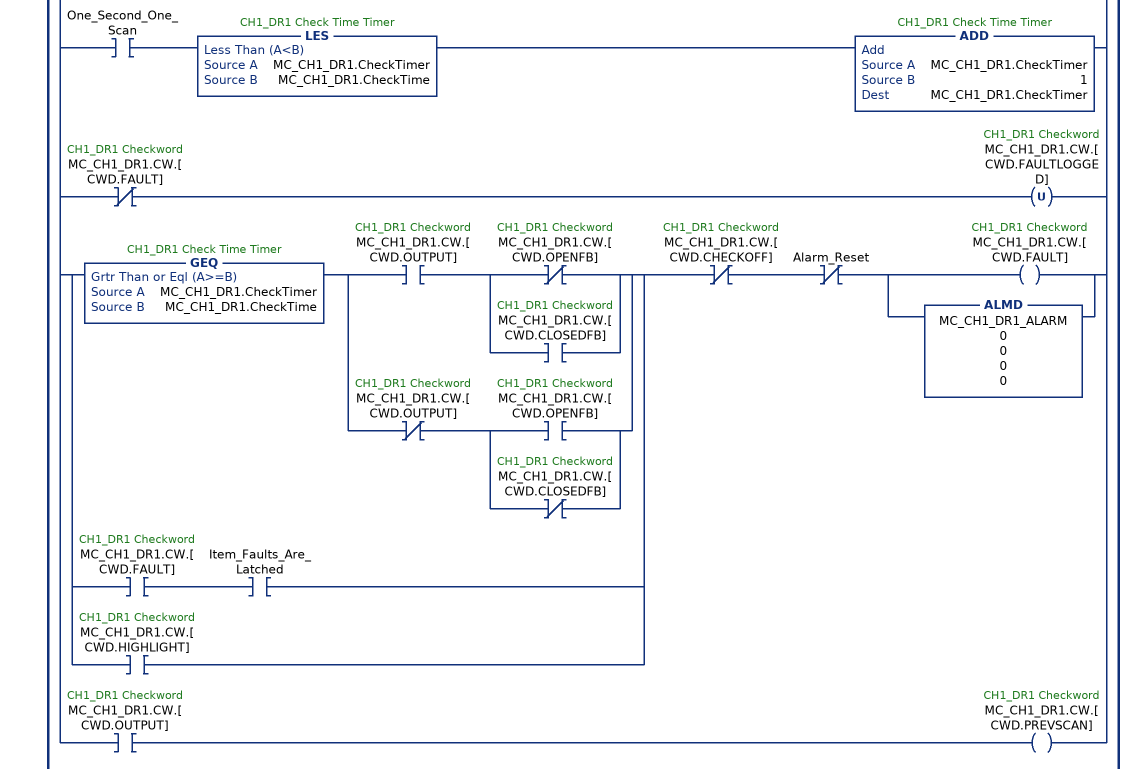
   14: [NEQ(MC_CH1_DR1.DriveBits,0) OTE(MC_CH1_DR1.CW.[CWD.AUTODRV]) ,[XIC(MC_CH1_DR1.CW.[CWD.AUTODRV]) XIO(MC_CH1_DR1.CW.[CWD.MANUAL]) ,XIC(MC_CH1_DR1.CW.[CWD.MANDRV]) XIC(MC_CH1_DR1.CW.[CWD.MANUAL]) ] OTE(MC_CH1_DR1.CW.[CWD.OUTPUT]) ,XIC(MC_CH1_DR1.CW.[CWD.OUTPUT]) OTE(MC_CH1_DR1_DR) ,XIC(S:FS) [OTU(MC_CH1_DR1.CW.[CWD.MANUAL]) ,LEQ(MC_CH1_DR1.CheckTime,0) MOV(Default_Check_Time,MC_CH1_DR1.CheckTime) ] ,[[XIC(MC_CH1_DR1_O) XIO(Item_Simulation_Flag) ,XIC(Item_Simulation_Flag) XIC(MC_CH1_DR1.CW.[CWD.OUTPUT]) XIO(MC_CH1_DR1.CW.[CWD.SIMFAIL]) ] OTE(MC_CH1_DR1.CW.[CWD.OPENFB]) ,[XIC(MC_CH1_DR1_C) XIO(Item_Simulation_Flag) ,XIC(Item_Simulation_Flag) XIO(MC_CH1_DR1.CW.[CWD.OUTPUT]) XIO(MC_CH1_DR1.CW.[CWD.SIMFAIL]) ] OTE(MC_CH1_DR1.CW.[CWD.CLOSEDFB]) ] ,[XIC(MC_CH1_DR1.CW.[CWD.OUTPUT]) XIO(MC_CH1_DR1.CW.[CWD.PREVSCAN]) ,XIO(MC_CH1_DR1.CW.[CWD.OUTPUT]) XIC(MC_CH1_DR1.CW.[CWD.PREVSCAN]) ] CLR(MC_CH1_DR1.CheckTimer) ,XIC(One_Second_One_Scan) LES(MC_CH1_DR1.CheckTimer,MC_CH1_DR1.CheckTime) ADD(MC_CH1_DR1.CheckTimer,1,MC_CH1_DR1.CheckTimer) ,XIO(MC_CH1_DR1.CW.[CWD.FAULT]) OTU(MC_CH1_DR1.CW.[CWD.FAULTLOGGED]) ,[GEQ(MC_CH1_DR1.CheckTimer,MC_CH1_DR1.CheckTime) [XIC(MC_CH1_DR1.CW.[CWD.OUTPUT]) [XIO(MC_CH1_DR1.CW.[CWD.OPENFB]) ,XIC(MC_CH1_DR1.CW.[CWD.CLOSEDFB]) ] ,XIO(MC_CH1_DR1.CW.[CWD.OUTPUT]) [XIC(MC_CH1_DR1.CW.[CWD.OPENFB]) ,XIO(MC_CH1_DR1.CW.[CWD.CLOSEDFB]) ] ] ,XIC(MC_CH1_DR1.CW.[CWD.FAULT]) XIC(Item_Faults_Are_Latched) ,XIC(MC_CH1_DR1.CW.[CWD.HIGHLIGHT]) ] XIO(MC_CH1_DR1.CW.[CWD.CHECKOFF]) XIO(Alarm_Reset) [OTE(MC_CH1_DR1.CW.[CWD.FAULT]) ,ALMD(MC_CH1_DR1_ALARM,0,0,0,0) ] ,XIC(MC_CH1_DR1.CW.[CWD.OUTPUT]) OTE(MC_CH1_DR1.CW.[CWD.PREVSCAN]) ];
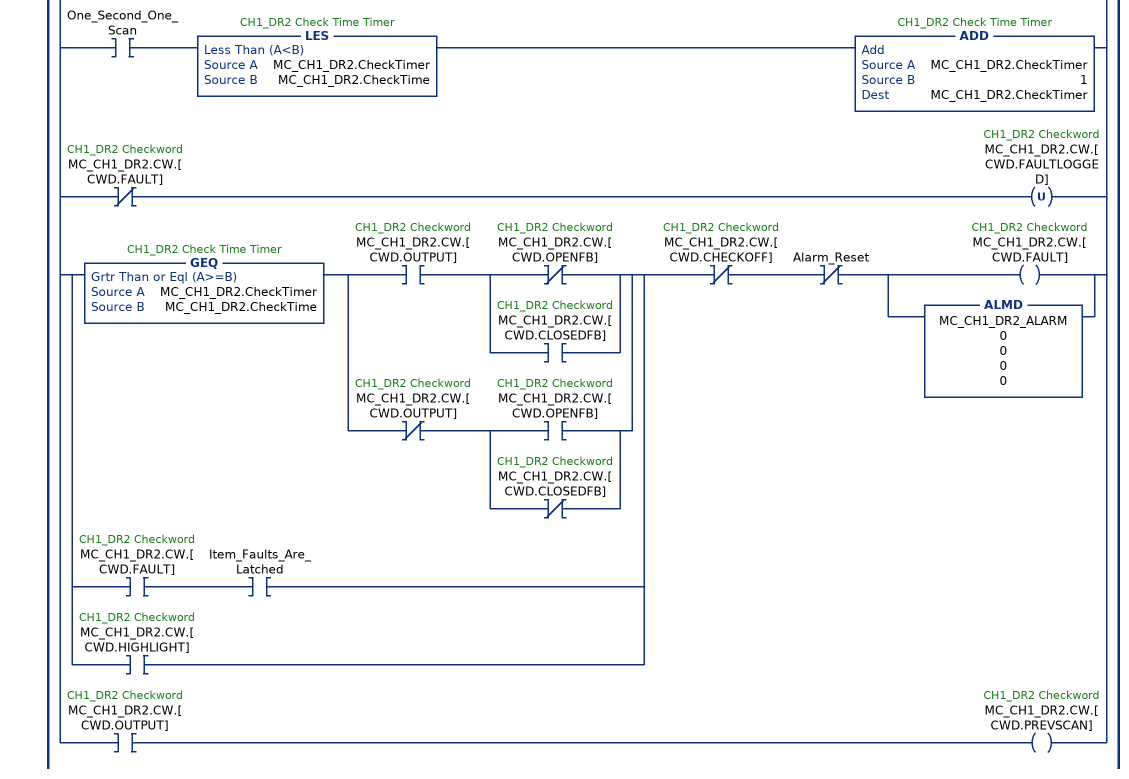
   15: [NEQ(MC_CH1_DR2.DriveBits,0) OTE(MC_CH1_DR2.CW.[CWD.AUTODRV]) ,[XIC(MC_CH1_DR2.CW.[CWD.AUTODRV]) XIO(MC_CH1_DR2.CW.[CWD.MANUAL]) ,XIC(MC_CH1_DR2.CW.[CWD.MANDRV]) XIC(MC_CH1_DR2.CW.[CWD.MANUAL]) ] OTE(MC_CH1_DR2.CW.[CWD.OUTPUT]) ,XIC(MC_CH1_DR2.CW.[CWD.OUTPUT]) OTE(MC_CH1_DR2_DR) ,XIC(S:FS) [OTU(MC_CH1_DR2.CW.[CWD.MANUAL]) ,LEQ(MC_CH1_DR2.CheckTime,0) MOV(Default_Check_Time,MC_CH1_DR2.CheckTime) ] ,[[XIC(MC_CH1_DR2_O) XIO(Item_Simulation_Flag) ,XIC(Item_Simulation_Flag) XIC(MC_CH1_DR2.CW.[CWD.OUTPUT]) XIO(MC_CH1_DR2.CW.[CWD.SIMFAIL]) ] OTE(MC_CH1_DR2.CW.[CWD.OPENFB]) ,[XIC(MC_CH1_DR2_C) XIO(Item_Simulation_Flag) ,XIC(Item_Simulation_Flag) XIO(MC_CH1_DR2.CW.[CWD.OUTPUT]) XIO(MC_CH1_DR2.CW.[CWD.SIMFAIL]) ] OTE(MC_CH1_DR2.CW.[CWD.CLOSEDFB]) ] ,[XIC(MC_CH1_DR2.CW.[CWD.OUTPUT]) XIO(MC_CH1_DR2.CW.[CWD.PREVSCAN]) ,XIO(MC_CH1_DR2.CW.[CWD.OUTPUT]) XIC(MC_CH1_DR2.CW.[CWD.PREVSCAN]) ] CLR(MC_CH1_DR2.CheckTimer) ,XIC(One_Second_One_Scan) LES(MC_CH1_DR2.CheckTimer,MC_CH1_DR2.CheckTime) ADD(MC_CH1_DR2.CheckTimer,1,MC_CH1_DR2.CheckTimer) ,XIO(MC_CH1_DR2.CW.[CWD.FAULT]) OTU(MC_CH1_DR2.CW.[CWD.FAULTLOGGED]) ,[GEQ(MC_CH1_DR2.CheckTimer,MC_CH1_DR2.CheckTime) [XIC(MC_CH1_DR2.CW.[CWD.OUTPUT]) [XIO(MC_CH1_DR2.CW.[CWD.OPENFB]) ,XIC(MC_CH1_DR2.CW.[CWD.CLOSEDFB]) ] ,XIO(MC_CH1_DR2.CW.[CWD.OUTPUT]) [XIC(MC_CH1_DR2.CW.[CWD.OPENFB]) ,XIO(MC_CH1_DR2.CW.[CWD.CLOSEDFB]) ] ] ,XIC(MC_CH1_DR2.CW.[CWD.FAULT]) XIC(Item_Faults_Are_Latched) ,XIC(MC_CH1_DR2.CW.[CWD.HIGHLIGHT]) ] XIO(MC_CH1_DR2.CW.[CWD.CHECKOFF]) XIO(Alarm_Reset) [OTE(MC_CH1_DR2.CW.[CWD.FAULT]) ,ALMD(MC_CH1_DR2_ALARM,0,0,0,0) ] ,XIC(MC_CH1_DR2.CW.[CWD.OUTPUT]) OTE(MC_CH1_DR2.CW.[CWD.PREVSCAN]) ];
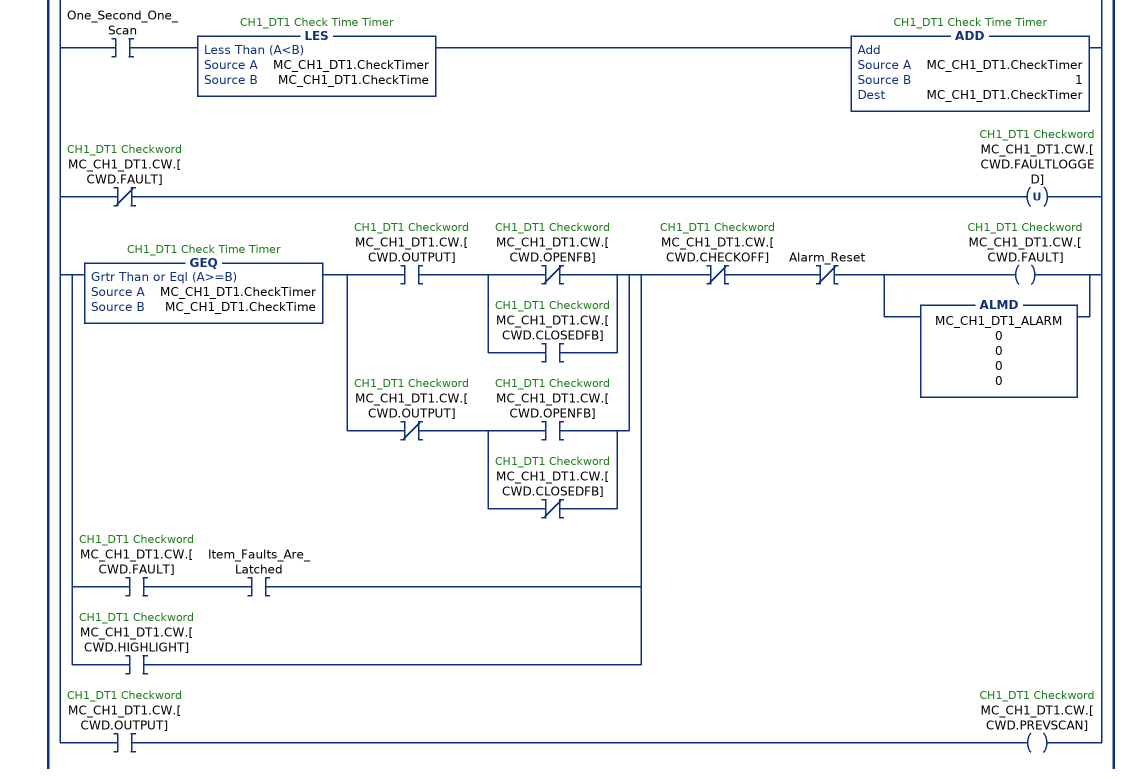
   16: [NEQ(MC_CH1_DT1.DriveBits,0) OTE(MC_CH1_DT1.CW.[CWD.AUTODRV]) ,[XIC(MC_CH1_DT1.CW.[CWD.AUTODRV]) XIO(MC_CH1_DT1.CW.[CWD.MANUAL]) ,XIC(MC_CH1_DT1.CW.[CWD.MANDRV]) XIC(MC_CH1_DT1.CW.[CWD.MANUAL]) ] OTE(MC_CH1_DT1.CW.[CWD.OUTPUT]) ,XIC(MC_CH1_DT1.CW.[CWD.OUTPUT]) OTE(MC_CH1_DT1_DR) ,XIC(S:FS) [OTU(MC_CH1_DT1.CW.[CWD.MANUAL]) ,LEQ(MC_CH1_DT1.CheckTime,0) MOV(Default_Check_Time,MC_CH1_DT1.CheckTime) ] ,[[XIC(MC_CH1_DT1_O) XIO(Item_Simulation_Flag) ,XIC(Item_Simulation_Flag) XIC(MC_CH1_DT1.CW.[CWD.OUTPUT]) XIO(MC_CH1_DT1.CW.[CWD.SIMFAIL]) ] OTE(MC_CH1_DT1.CW.[CWD.OPENFB]) ,[XIC(MC_CH1_DT1_C) XIO(Item_Simulation_Flag) ,XIC(Item_Simulation_Flag) XIO(MC_CH1_DT1.CW.[CWD.OUTPUT]) XIO(MC_CH1_DT1.CW.[CWD.SIMFAIL]) ] OTE(MC_CH1_DT1.CW.[CWD.CLOSEDFB]) ] ,[XIC(MC_CH1_DT1.CW.[CWD.OUTPUT]) XIO(MC_CH1_DT1.CW.[CWD.PREVSCAN]) ,XIO(MC_CH1_DT1.CW.[CWD.OUTPUT]) XIC(MC_CH1_DT1.CW.[CWD.PREVSCAN]) ] CLR(MC_CH1_DT1.CheckTimer) ,XIC(One_Second_One_Scan) LES(MC_CH1_DT1.CheckTimer,MC_CH1_DT1.CheckTime) ADD(MC_CH1_DT1.CheckTimer,1,MC_CH1_DT1.CheckTimer) ,XIO(MC_CH1_DT1.CW.[CWD.FAULT]) OTU(MC_CH1_DT1.CW.[CWD.FAULTLOGGED]) ,[GEQ(MC_CH1_DT1.CheckTimer,MC_CH1_DT1.CheckTime) [XIC(MC_CH1_DT1.CW.[CWD.OUTPUT]) [XIO(MC_CH1_DT1.CW.[CWD.OPENFB]) ,XIC(MC_CH1_DT1.CW.[CWD.CLOSEDFB]) ] ,XIO(MC_CH1_DT1.CW.[CWD.OUTPUT]) [XIC(MC_CH1_DT1.CW.[CWD.OPENFB]) ,XIO(MC_CH1_DT1.CW.[CWD.CLOSEDFB]) ] ] ,XIC(MC_CH1_DT1.CW.[CWD.FAULT]) XIC(Item_Faults_Are_Latched) ,XIC(MC_CH1_DT1.CW.[CWD.HIGHLIGHT]) ] XIO(MC_CH1_DT1.CW.[CWD.CHECKOFF]) XIO(Alarm_Reset) [OTE(MC_CH1_DT1.CW.[CWD.FAULT]) ,ALMD(MC_CH1_DT1_ALARM,0,0,0,0) ] ,XIC(MC_CH1_DT1.CW.[CWD.OUTPUT]) OTE(MC_CH1_DT1.CW.[CWD.PREVSCAN]) ];
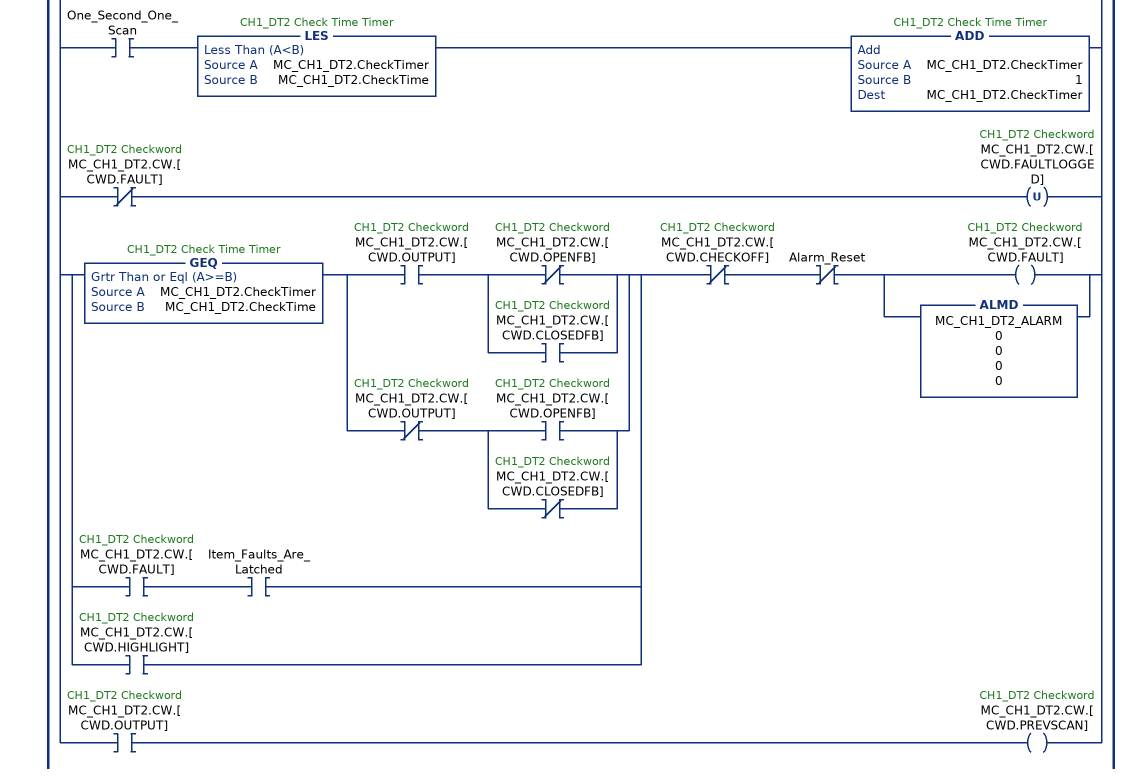
   17: [NEQ(MC_CH1_DT2.DriveBits,0) OTE(MC_CH1_DT2.CW.[CWD.AUTODRV]) ,[XIC(MC_CH1_DT2.CW.[CWD.AUTODRV]) XIO(MC_CH1_DT2.CW.[CWD.MANUAL]) ,XIC(MC_CH1_DT2.CW.[CWD.MANDRV]) XIC(MC_CH1_DT2.CW.[CWD.MANUAL]) ] OTE(MC_CH1_DT2.CW.[CWD.OUTPUT]) ,XIC(MC_CH1_DT2.CW.[CWD.OUTPUT]) OTE(MC_CH1_DT2_DR) ,XIC(S:FS) [OTU(MC_CH1_DT2.CW.[CWD.MANUAL]) ,LEQ(MC_CH1_DT2.CheckTime,0) MOV(Default_Check_Time,MC_CH1_DT2.CheckTime) ] ,[[XIC(MC_CH1_DT2_O) XIO(Item_Simulation_Flag) ,XIC(Item_Simulation_Flag) XIC(MC_CH1_DT2.CW.[CWD.OUTPUT]) XIO(MC_CH1_DT2.CW.[CWD.SIMFAIL]) ] OTE(MC_CH1_DT2.CW.[CWD.OPENFB]) ,[XIC(MC_CH1_DT2_C) XIO(Item_Simulation_Flag) ,XIC(Item_Simulation_Flag) XIO(MC_CH1_DT2.CW.[CWD.OUTPUT]) XIO(MC_CH1_DT2.CW.[CWD.SIMFAIL]) ] OTE(MC_CH1_DT2.CW.[CWD.CLOSEDFB]) ] ,[XIC(MC_CH1_DT2.CW.[CWD.OUTPUT]) XIO(MC_CH1_DT2.CW.[CWD.PREVSCAN]) ,XIO(MC_CH1_DT2.CW.[CWD.OUTPUT]) XIC(MC_CH1_DT2.CW.[CWD.PREVSCAN]) ] CLR(MC_CH1_DT2.CheckTimer) ,XIC(One_Second_One_Scan) LES(MC_CH1_DT2.CheckTimer,MC_CH1_DT2.CheckTime) ADD(MC_CH1_DT2.CheckTimer,1,MC_CH1_DT2.CheckTimer) ,XIO(MC_CH1_DT2.CW.[CWD.FAULT]) OTU(MC_CH1_DT2.CW.[CWD.FAULTLOGGED]) ,[GEQ(MC_CH1_DT2.CheckTimer,MC_CH1_DT2.CheckTime) [XIC(MC_CH1_DT2.CW.[CWD.OUTPUT]) [XIO(MC_CH1_DT2.CW.[CWD.OPENFB]) ,XIC(MC_CH1_DT2.CW.[CWD.CLOSEDFB]) ] ,XIO(MC_CH1_DT2.CW.[CWD.OUTPUT]) [XIC(MC_CH1_DT2.CW.[CWD.OPENFB]) ,XIO(MC_CH1_DT2.CW.[CWD.CLOSEDFB]) ] ] ,XIC(MC_CH1_DT2.CW.[CWD.FAULT]) XIC(Item_Faults_Are_Latched) ,XIC(MC_CH1_DT2.CW.[CWD.HIGHLIGHT]) ] XIO(MC_CH1_DT2.CW.[CWD.CHECKOFF]) XIO(Alarm_Reset) [OTE(MC_CH1_DT2.CW.[CWD.FAULT]) ,ALMD(MC_CH1_DT2_ALARM,0,0,0,0) ] ,XIC(MC_CH1_DT2.CW.[CWD.OUTPUT]) OTE(MC_CH1_DT2.CW.[CWD.PREVSCAN]) ];
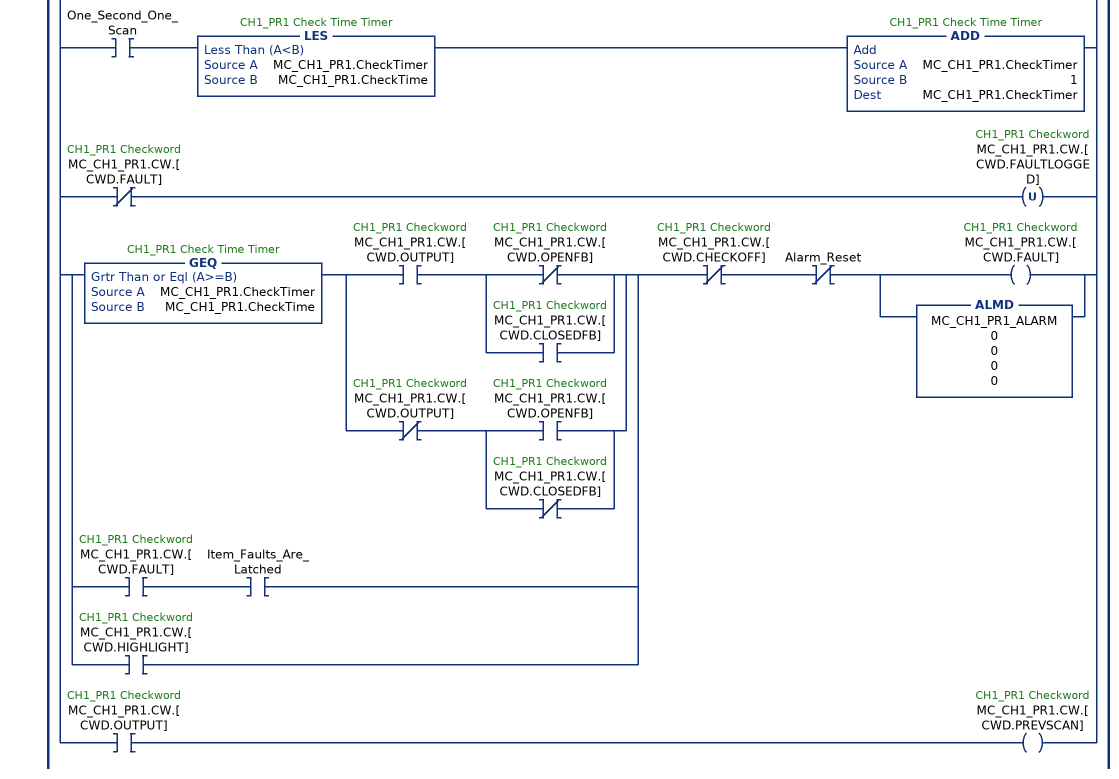
   18: [NEQ(MC_CH1_PR1.DriveBits,0) OTE(MC_CH1_PR1.CW.[CWD.AUTODRV]) ,[XIC(MC_CH1_PR1.CW.[CWD.AUTODRV]) XIO(MC_CH1_PR1.CW.[CWD.MANUAL]) ,XIC(MC_CH1_PR1.CW.[CWD.MANDRV]) XIC(MC_CH1_PR1.CW.[CWD.MANUAL]) ] OTE(MC_CH1_PR1.CW.[CWD.OUTPUT]) ,XIC(MC_CH1_PR1.CW.[CWD.OUTPUT]) OTE(MC_CH1_PR1_DR) ,XIC(S:FS) [OTU(MC_CH1_PR1.CW.[CWD.MANUAL]) ,LEQ(MC_CH1_PR1.CheckTime,0) MOV(Default_Check_Time,MC_CH1_PR1.CheckTime) ] ,[[XIC(MC_CH1_PR1_O) XIO(Item_Simulation_Flag) ,XIC(Item_Simulation_Flag) XIC(MC_CH1_PR1.CW.[CWD.OUTPUT]) XIO(MC_CH1_PR1.CW.[CWD.SIMFAIL]) ] OTE(MC_CH1_PR1.CW.[CWD.OPENFB]) ,[XIC(MC_CH1_PR1_C) XIO(Item_Simulation_Flag) ,XIC(Item_Simulation_Flag) XIO(MC_CH1_PR1.CW.[CWD.OUTPUT]) XIO(MC_CH1_PR1.CW.[CWD.SIMFAIL]) ] OTE(MC_CH1_PR1.CW.[CWD.CLOSEDFB]) ] ,[XIC(MC_CH1_PR1.CW.[CWD.OUTPUT]) XIO(MC_CH1_PR1.CW.[CWD.PREVSCAN]) ,XIO(MC_CH1_PR1.CW.[CWD.OUTPUT]) XIC(MC_CH1_PR1.CW.[CWD.PREVSCAN]) ] CLR(MC_CH1_PR1.CheckTimer) ,XIC(One_Second_One_Scan) LES(MC_CH1_PR1.CheckTimer,MC_CH1_PR1.CheckTime) ADD(MC_CH1_PR1.CheckTimer,1,MC_CH1_PR1.CheckTimer) ,XIO(MC_CH1_PR1.CW.[CWD.FAULT]) OTU(MC_CH1_PR1.CW.[CWD.FAULTLOGGED]) ,[GEQ(MC_CH1_PR1.CheckTimer,MC_CH1_PR1.CheckTime) [XIC(MC_CH1_PR1.CW.[CWD.OUTPUT]) [XIO(MC_CH1_PR1.CW.[CWD.OPENFB]) ,XIC(MC_CH1_PR1.CW.[CWD.CLOSEDFB]) ] ,XIO(MC_CH1_PR1.CW.[CWD.OUTPUT]) [XIC(MC_CH1_PR1.CW.[CWD.OPENFB]) ,XIO(MC_CH1_PR1.CW.[CWD.CLOSEDFB]) ] ] ,XIC(MC_CH1_PR1.CW.[CWD.FAULT]) XIC(Item_Faults_Are_Latched) ,XIC(MC_CH1_PR1.CW.[CWD.HIGHLIGHT]) ] XIO(MC_CH1_PR1.CW.[CWD.CHECKOFF]) XIO(Alarm_Reset) [OTE(MC_CH1_PR1.CW.[CWD.FAULT]) ,ALMD(MC_CH1_PR1_ALARM,0,0,0,0) ] ,XIC(MC_CH1_PR1.CW.[CWD.OUTPUT]) OTE(MC_CH1_PR1.CW.[CWD.PREVSCAN]) ];
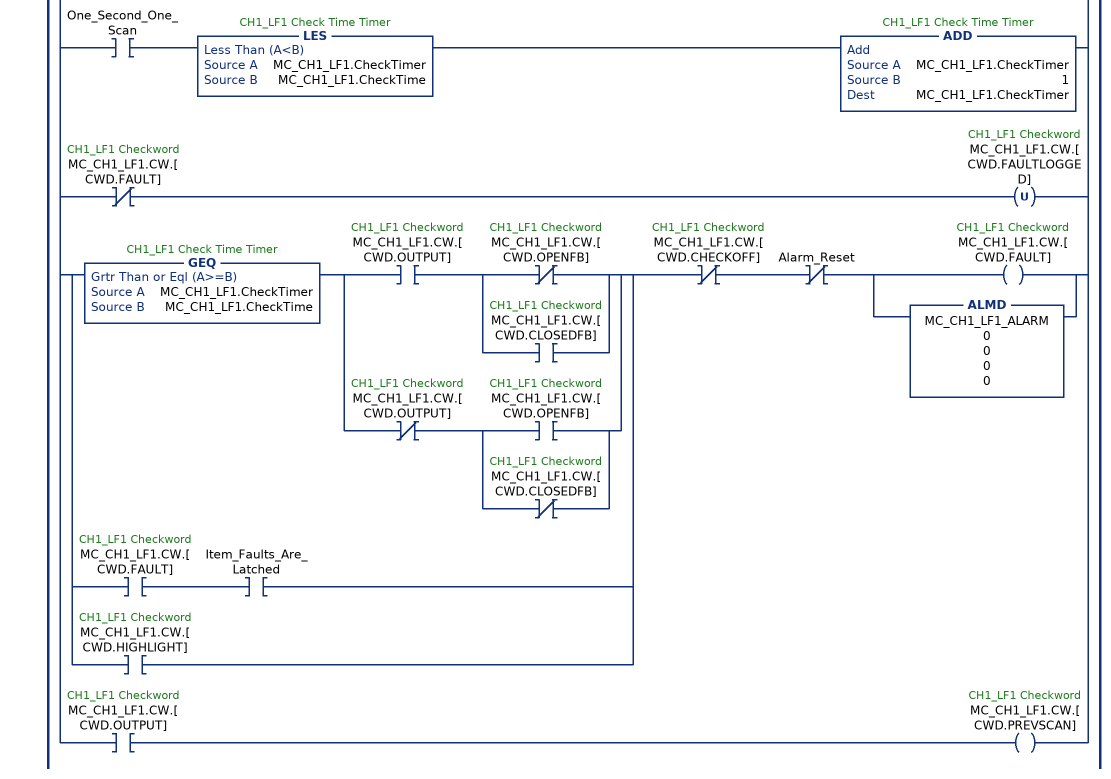
   19: [NEQ(MC_CH1_LF1.DriveBits,0) OTE(MC_CH1_LF1.CW.[CWD.AUTODRV]) ,[XIC(MC_CH1_LF1.CW.[CWD.AUTODRV]) XIO(MC_CH1_LF1.CW.[CWD.MANUAL]) ,XIC(MC_CH1_LF1.CW.[CWD.MANDRV]) XIC(MC_CH1_LF1.CW.[CWD.MANUAL]) ] OTE(MC_CH1_LF1.CW.[CWD.OUTPUT]) ,XIC(MC_CH1_LF1.CW.[CWD.OUTPUT]) OTE(MC_CH1_LF1_DR) ,XIC(S:FS) [OTU(MC_CH1_LF1.CW.[CWD.MANUAL]) ,LEQ(MC_CH1_LF1.CheckTime,0) MOV(Default_Check_Time,MC_CH1_LF1.CheckTime) ] ,[[XIC(MC_CH1_LF1_O) XIO(Item_Simulation_Flag) ,XIC(Item_Simulation_Flag) XIC(MC_CH1_LF1.CW.[CWD.OUTPUT]) XIO(MC_CH1_LF1.CW.[CWD.SIMFAIL]) ] OTE(MC_CH1_LF1.CW.[CWD.OPENFB]) ,[XIC(MC_CH1_LF1_C) XIO(Item_Simulation_Flag) ,XIC(Item_Simulation_Flag) XIO(MC_CH1_LF1.CW.[CWD.OUTPUT]) XIO(MC_CH1_LF1.CW.[CWD.SIMFAIL]) ] OTE(MC_CH1_LF1.CW.[CWD.CLOSEDFB]) ] ,[XIC(MC_CH1_LF1.CW.[CWD.OUTPUT]) XIO(MC_CH1_LF1.CW.[CWD.PREVSCAN]) ,XIO(MC_CH1_LF1.CW.[CWD.OUTPUT]) XIC(MC_CH1_LF1.CW.[CWD.PREVSCAN]) ] CLR(MC_CH1_LF1.CheckTimer) ,XIC(One_Second_One_Scan) LES(MC_CH1_LF1.CheckTimer,MC_CH1_LF1.CheckTime) ADD(MC_CH1_LF1.CheckTimer,1,MC_CH1_LF1.CheckTimer) ,XIO(MC_CH1_LF1.CW.[CWD.FAULT]) OTU(MC_CH1_LF1.CW.[CWD.FAULTLOGGED]) ,[GEQ(MC_CH1_LF1.CheckTimer,MC_CH1_LF1.CheckTime) [XIC(MC_CH1_LF1.CW.[CWD.OUTPUT]) [XIO(MC_CH1_LF1.CW.[CWD.OPENFB]) ,XIC(MC_CH1_LF1.CW.[CWD.CLOSEDFB]) ] ,XIO(MC_CH1_LF1.CW.[CWD.OUTPUT]) [XIC(MC_CH1_LF1.CW.[CWD.OPENFB]) ,XIO(MC_CH1_LF1.CW.[CWD.CLOSEDFB]) ] ] ,XIC(MC_CH1_LF1.CW.[CWD.FAULT]) XIC(Item_Faults_Are_Latched) ,XIC(MC_CH1_LF1.CW.[CWD.HIGHLIGHT]) ] XIO(MC_CH1_LF1.CW.[CWD.CHECKOFF]) XIO(Alarm_Reset) [OTE(MC_CH1_LF1.CW.[CWD.FAULT]) ,ALMD(MC_CH1_LF1_ALARM,0,0,0,0) ] ,XIC(MC_CH1_LF1.CW.[CWD.OUTPUT]) OTE(MC_CH1_LF1.CW.[CWD.PREVSCAN]) ];
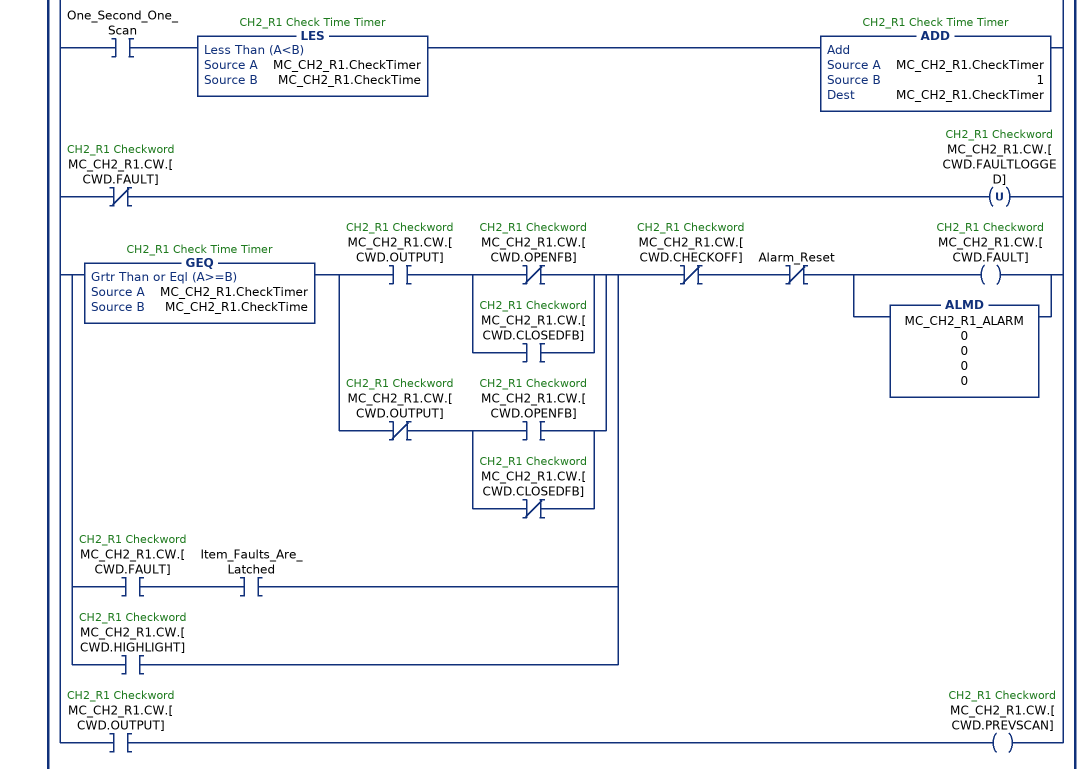
   20: [NEQ(MC_CH2_R1.DriveBits,0) OTE(MC_CH2_R1.CW.[CWD.AUTODRV]) ,[XIC(MC_CH2_R1.CW.[CWD.AUTODRV]) XIO(MC_CH2_R1.CW.[CWD.MANUAL]) ,XIC(MC_CH2_R1.CW.[CWD.MANDRV]) XIC(MC_CH2_R1.CW.[CWD.MANUAL]) ] OTE(MC_CH2_R1.CW.[CWD.OUTPUT]) ,XIC(MC_CH2_R1.CW.[CWD.OUTPUT]) OTE(MC_CH2_R1_DR) ,XIC(S:FS) [OTU(MC_CH2_R1.CW.[CWD.MANUAL]) ,LEQ(MC_CH2_R1.CheckTime,0) MOV(Default_Check_Time,MC_CH2_R1.CheckTime) ] ,[[XIC(MC_CH2_R1_O) XIO(Item_Simulation_Flag) ,XIC(Item_Simulation_Flag) XIC(MC_CH2_R1.CW.[CWD.OUTPUT]) XIO(MC_CH2_R1.CW.[CWD.SIMFAIL]) ] OTE(MC_CH2_R1.CW.[CWD.OPENFB]) ,[XIC(MC_CH2_R1_C) XIO(Item_Simulation_Flag) ,XIC(Item_Simulation_Flag) XIO(MC_CH2_R1.CW.[CWD.OUTPUT]) XIO(MC_CH2_R1.CW.[CWD.SIMFAIL]) ] OTE(MC_CH2_R1.CW.[CWD.CLOSEDFB]) ] ,[XIC(MC_CH2_R1.CW.[CWD.OUTPUT]) XIO(MC_CH2_R1.CW.[CWD.PREVSCAN]) ,XIO(MC_CH2_R1.CW.[CWD.OUTPUT]) XIC(MC_CH2_R1.CW.[CWD.PREVSCAN]) ] CLR(MC_CH2_R1.CheckTimer) ,XIC(One_Second_One_Scan) LES(MC_CH2_R1.CheckTimer,MC_CH2_R1.CheckTime) ADD(MC_CH2_R1.CheckTimer,1,MC_CH2_R1.CheckTimer) ,XIO(MC_CH2_R1.CW.[CWD.FAULT]) OTU(MC_CH2_R1.CW.[CWD.FAULTLOGGED]) ,[GEQ(MC_CH2_R1.CheckTimer,MC_CH2_R1.CheckTime) [XIC(MC_CH2_R1.CW.[CWD.OUTPUT]) [XIO(MC_CH2_R1.CW.[CWD.OPENFB]) ,XIC(MC_CH2_R1.CW.[CWD.CLOSEDFB]) ] ,XIO(MC_CH2_R1.CW.[CWD.OUTPUT]) [XIC(MC_CH2_R1.CW.[CWD.OPENFB]) ,XIO(MC_CH2_R1.CW.[CWD.CLOSEDFB]) ] ] ,XIC(MC_CH2_R1.CW.[CWD.FAULT]) XIC(Item_Faults_Are_Latched) ,XIC(MC_CH2_R1.CW.[CWD.HIGHLIGHT]) ] XIO(MC_CH2_R1.CW.[CWD.CHECKOFF]) XIO(Alarm_Reset) [OTE(MC_CH2_R1.CW.[CWD.FAULT]) ,ALMD(MC_CH2_R1_ALARM,0,0,0,0) ] ,XIC(MC_CH2_R1.CW.[CWD.OUTPUT]) OTE(MC_CH2_R1.CW.[CWD.PREVSCAN]) ];
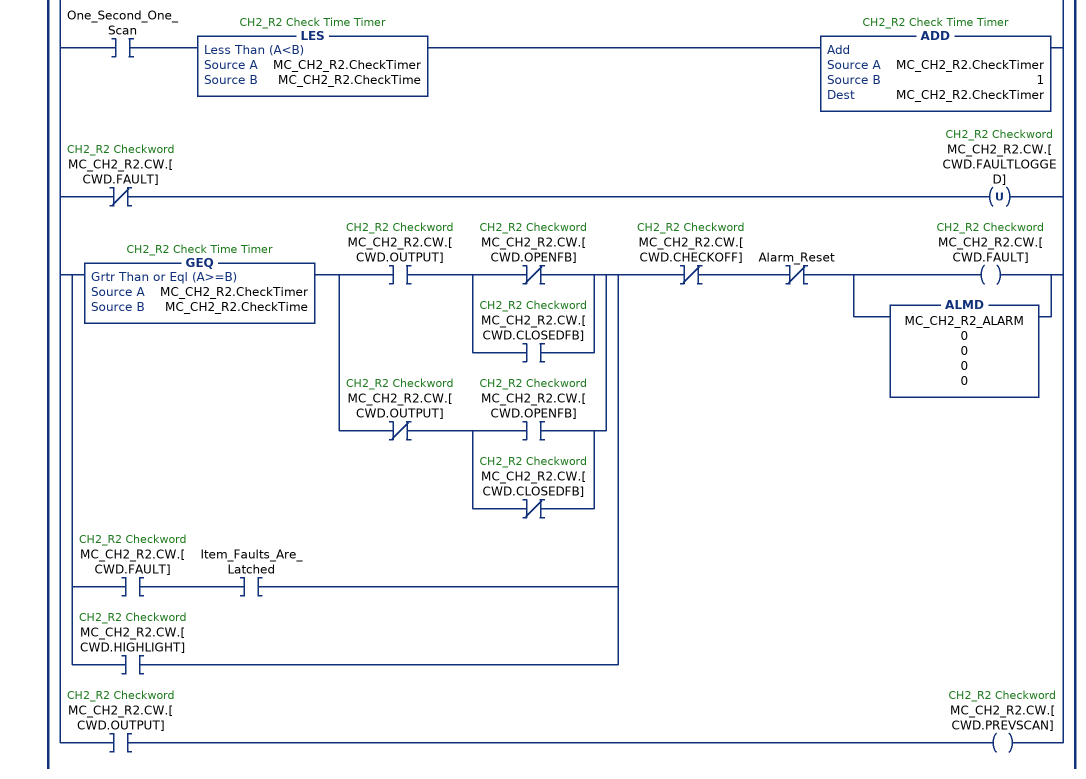
   21: [NEQ(MC_CH2_R2.DriveBits,0) OTE(MC_CH2_R2.CW.[CWD.AUTODRV]) ,[XIC(MC_CH2_R2.CW.[CWD.AUTODRV]) XIO(MC_CH2_R2.CW.[CWD.MANUAL]) ,XIC(MC_CH2_R2.CW.[CWD.MANDRV]) XIC(MC_CH2_R2.CW.[CWD.MANUAL]) ] OTE(MC_CH2_R2.CW.[CWD.OUTPUT]) ,XIC(MC_CH2_R2.CW.[CWD.OUTPUT]) OTE(MC_CH2_R2_DR) ,XIC(S:FS) [OTU(MC_CH2_R2.CW.[CWD.MANUAL]) ,LEQ(MC_CH2_R2.CheckTime,0) MOV(Default_Check_Time,MC_CH2_R2.CheckTime) ] ,[[XIC(MC_CH2_R2_O) XIO(Item_Simulation_Flag) ,XIC(Item_Simulation_Flag) XIC(MC_CH2_R2.CW.[CWD.OUTPUT]) XIO(MC_CH2_R2.CW.[CWD.SIMFAIL]) ] OTE(MC_CH2_R2.CW.[CWD.OPENFB]) ,[XIC(MC_CH2_R2_C) XIO(Item_Simulation_Flag) ,XIC(Item_Simulation_Flag) XIO(MC_CH2_R2.CW.[CWD.OUTPUT]) XIO(MC_CH2_R2.CW.[CWD.SIMFAIL]) ] OTE(MC_CH2_R2.CW.[CWD.CLOSEDFB]) ] ,[XIC(MC_CH2_R2.CW.[CWD.OUTPUT]) XIO(MC_CH2_R2.CW.[CWD.PREVSCAN]) ,XIO(MC_CH2_R2.CW.[CWD.OUTPUT]) XIC(MC_CH2_R2.CW.[CWD.PREVSCAN]) ] CLR(MC_CH2_R2.CheckTimer) ,XIC(One_Second_One_Scan) LES(MC_CH2_R2.CheckTimer,MC_CH2_R2.CheckTime) ADD(MC_CH2_R2.CheckTimer,1,MC_CH2_R2.CheckTimer) ,XIO(MC_CH2_R2.CW.[CWD.FAULT]) OTU(MC_CH2_R2.CW.[CWD.FAULTLOGGED]) ,[GEQ(MC_CH2_R2.CheckTimer,MC_CH2_R2.CheckTime) [XIC(MC_CH2_R2.CW.[CWD.OUTPUT]) [XIO(MC_CH2_R2.CW.[CWD.OPENFB]) ,XIC(MC_CH2_R2.CW.[CWD.CLOSEDFB]) ] ,XIO(MC_CH2_R2.CW.[CWD.OUTPUT]) [XIC(MC_CH2_R2.CW.[CWD.OPENFB]) ,XIO(MC_CH2_R2.CW.[CWD.CLOSEDFB]) ] ] ,XIC(MC_CH2_R2.CW.[CWD.FAULT]) XIC(Item_Faults_Are_Latched) ,XIC(MC_CH2_R2.CW.[CWD.HIGHLIGHT]) ] XIO(MC_CH2_R2.CW.[CWD.CHECKOFF]) XIO(Alarm_Reset) [OTE(MC_CH2_R2.CW.[CWD.FAULT]) ,ALMD(MC_CH2_R2_ALARM,0,0,0,0) ] ,XIC(MC_CH2_R2.CW.[CWD.OUTPUT]) OTE(MC_CH2_R2.CW.[CWD.PREVSCAN]) ];
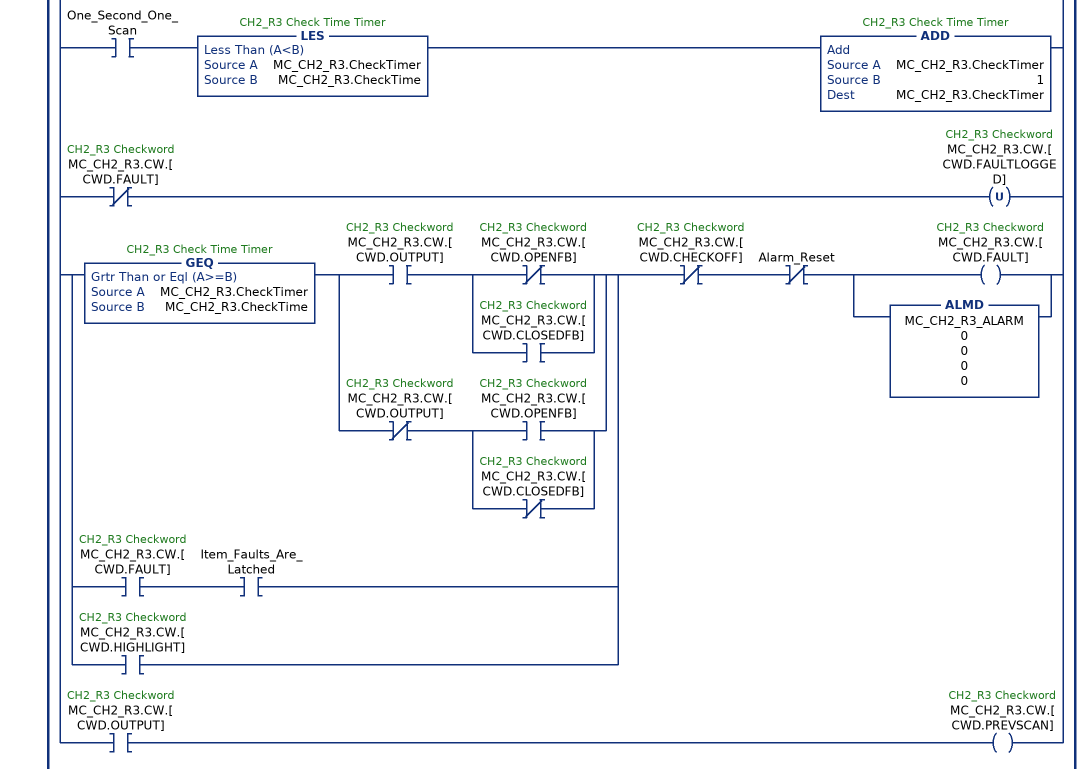
   22: [NEQ(MC_CH2_R3.DriveBits,0) OTE(MC_CH2_R3.CW.[CWD.AUTODRV]) ,[XIC(MC_CH2_R3.CW.[CWD.AUTODRV]) XIO(MC_CH2_R3.CW.[CWD.MANUAL]) ,XIC(MC_CH2_R3.CW.[CWD.MANDRV]) XIC(MC_CH2_R3.CW.[CWD.MANUAL]) ] OTE(MC_CH2_R3.CW.[CWD.OUTPUT]) ,XIC(MC_CH2_R3.CW.[CWD.OUTPUT]) OTE(MC_CH2_R3_DR) ,XIC(S:FS) [OTU(MC_CH2_R3.CW.[CWD.MANUAL]) ,LEQ(MC_CH2_R3.CheckTime,0) MOV(Default_Check_Time,MC_CH2_R3.CheckTime) ] ,[[XIC(MC_CH2_R3_O) XIO(Item_Simulation_Flag) ,XIC(Item_Simulation_Flag) XIC(MC_CH2_R3.CW.[CWD.OUTPUT]) XIO(MC_CH2_R3.CW.[CWD.SIMFAIL]) ] OTE(MC_CH2_R3.CW.[CWD.OPENFB]) ,[XIC(MC_CH2_R3_C) XIO(Item_Simulation_Flag) ,XIC(Item_Simulation_Flag) XIO(MC_CH2_R3.CW.[CWD.OUTPUT]) XIO(MC_CH2_R3.CW.[CWD.SIMFAIL]) ] OTE(MC_CH2_R3.CW.[CWD.CLOSEDFB]) ] ,[XIC(MC_CH2_R3.CW.[CWD.OUTPUT]) XIO(MC_CH2_R3.CW.[CWD.PREVSCAN]) ,XIO(MC_CH2_R3.CW.[CWD.OUTPUT]) XIC(MC_CH2_R3.CW.[CWD.PREVSCAN]) ] CLR(MC_CH2_R3.CheckTimer) ,XIC(One_Second_One_Scan) LES(MC_CH2_R3.CheckTimer,MC_CH2_R3.CheckTime) ADD(MC_CH2_R3.CheckTimer,1,MC_CH2_R3.CheckTimer) ,XIO(MC_CH2_R3.CW.[CWD.FAULT]) OTU(MC_CH2_R3.CW.[CWD.FAULTLOGGED]) ,[GEQ(MC_CH2_R3.CheckTimer,MC_CH2_R3.CheckTime) [XIC(MC_CH2_R3.CW.[CWD.OUTPUT]) [XIO(MC_CH2_R3.CW.[CWD.OPENFB]) ,XIC(MC_CH2_R3.CW.[CWD.CLOSEDFB]) ] ,XIO(MC_CH2_R3.CW.[CWD.OUTPUT]) [XIC(MC_CH2_R3.CW.[CWD.OPENFB]) ,XIO(MC_CH2_R3.CW.[CWD.CLOSEDFB]) ] ] ,XIC(MC_CH2_R3.CW.[CWD.FAULT]) XIC(Item_Faults_Are_Latched) ,XIC(MC_CH2_R3.CW.[CWD.HIGHLIGHT]) ] XIO(MC_CH2_R3.CW.[CWD.CHECKOFF]) XIO(Alarm_Reset) [OTE(MC_CH2_R3.CW.[CWD.FAULT]) ,ALMD(MC_CH2_R3_ALARM,0,0,0,0) ] ,XIC(MC_CH2_R3.CW.[CWD.OUTPUT]) OTE(MC_CH2_R3.CW.[CWD.PREVSCAN]) ];